               x10 : Bool;   // Direct output 1 via traversing block
               x11 : Bool;   // Direct output 2 via traversing block
               x12 : Bool;   // Fixed stop reached
               x13 : Bool;   // Fixed stop clamping torque reached
               x14 : Bool;   // Travel to fixed stop active
               x15 : Bool;   // Traversing command active
               x0 : Bool;   // Tracking mode active
               x1 : Bool;   // Velocity limit active
               x2 : Bool;   // Setpoint available
               x3 : Bool;   // Printing mark outside outer window
               x4 : Bool;   // Axis moves forwards
               x5 : Bool;   // Axis moves backwards
               x6 : Bool;   // Software limit switch minus reached
               x7 : Bool;   // Software limit switch plus reached
            END_STRUCT;
            dFDB_TARGET : DInt;   // R2060[5].Feedback target
            dXIST_A : DInt;   // R2521[0].Actual position value
            dNIST_B : DInt;   // R63.Actual speed value
            iFAULT_CODE : Int;   // R2131.Actual fault code
            iWARN_CODE : Int;   // R2132.Actual alarm code
            iUser : Int;
         END_STRUCT;
         tW : Struct   // WRITE
            tSTW1 : Struct   // CONTROL WORD 1
               x8 : Bool;   // P2589.EPOS jog 1 signal source
               x9 : Bool;   // P2590.EPOS jog 2 signal source
               x10 : Bool;   // P854[0].Control by PLC
               x11 : Bool;   // P2595.EPOS referencing start
               x12 : Bool;   // Reserved
               x13 : Bool;   // P2633.EPOS external block change
               x14 : Bool;   // Reserved
               x15 : Bool;   // P855[0] Brake release
               x0 : Bool;   // P840[0].ON/OFF
               x1 : Bool;   // P844[0].OFF2
               x2 : Bool;   // P848[0].OFF3
               x3 : Bool;   // P852[0].Enable operation
               x4 : Bool;   // P2641.EPOS abort traversing task
               x5 : Bool;   // P2640.EPOS intermediate STOP
               x6 : Bool;   // P2631.EPOS activate traversing task
               x7 : Bool;   // P2103.Acknowledge faults
            END_STRUCT;
            tPOS_STW1 : Struct   // POSITIONER CONTROL WORD 2
               x8 : Bool;   // P2648.EPOS direct setpoint input/MDI positioning type
               x9 : Bool;   // P2651.EPOS direct setpoint input/MDI direction selection positive
               x10 : Bool;   // P2652.EPOS direct setpoint input/MDI direction selection negative
               x11 : Bool;   // Reserved
               x12 : Bool;   // P2649.EPOS direct setpoint input/MDI transfer type selection
               x13 : Bool;   // Reserved
               x14 : Bool;   // P2653.EPOS direct setpoint input/MDI setting-up selection
               x15 : Bool;   // P2647.EPOS direct setpoint input/MDI selection
               x0 : Bool;   // P2525.EPOS traversing block selection, bit 0
               x1 : Bool;   // P2526.EPOS traversing block selection, bit 1
               x2 : Bool;   // P2527.EPOS traversing block selection, bit 2
               x3 : Bool;   // P2528.EPOS traversing block selection, bit 3
               x4 : Bool;   // P2529.EPOS traversing block selection, bit 4
               x5 : Bool;   // P2530.EPOS traversing block selection, bit 5
               x6 : Bool;   // Reserved
               x7 : Bool;   // Reserved
            END_STRUCT;
            tPOS_STW2 : Struct   // POSITIONER CONTROL WORD 3
               x8 : Bool;   // P2597.EPOS referencing type selection
               x9 : Bool;   // P2604.EPOS search for reference, start direction
               x10 : Bool;   // P2510.LR selecting measuring probe evaluation
               x11 : Bool;   // P2511.LR measuring probe evaluation edge
               x12 : Bool;   // Reserved
               x13 : Bool;   // Reserved
               x14 : Bool;   // P2582.EPOS software limit switch activation
               x15 : Bool;   // P2568.EPOS STOP cam activation
               x0 : Bool;   // P2655.EPOS select tracking mode
               x1 : Bool;   // P2596.EPOS set reference point
               x2 : Bool;   // P2612.EPOS search for reference cam
               x3 : Bool;   // Reserved
               x4 : Bool;   // Reserved
               x5 : Bool;   // P2591.EPOS jogging incremental
               x6 : Bool;   // Reserved
               x7 : Bool;   // Reserved
            END_STRUCT;
            iSTW2 : Int;   // P2045.CONTROL WORD 4
            iOVERRIDE : Int;   // P2646.Override % [0-16384]
            dMDI_TARPOS : DInt;   // P2642.Target position for MDI
            dMDI_VELOCITY : DInt;   // P2643.Speed reference for MDI
            iMDI_ACC : Int;   // P2644.Acceleration ramp % for MDI [0-16384]
            iMDI_DEC : Int;   // P2645.Deceleration ramp % for MDI [0-16384]
            iUser : Int;
         END_STRUCT;
      END_STRUCT;
   END_VAR
   VAR_TEMP
      TMP_dOldValue_AR1 : DInt;
      TMP_dOldValue_AR2 : DInt;
      TMP_x : Bool;
      TMP_i : Int;
      TMP_d : DInt;
      TMP_r : Real;
      TMP_a : ANY;
      TMP_dZero : DInt;
      TMP_xAlwaysON : Bool;
      TMP_rActualSpeed : Real;
      TMP_iAddressLength : Int;
      TMP_iRetVal : Int;
      TMP_dActualPosFiltered_cdeg : DInt;   // Actual position filtered [°/100]
      TMP_dActualPosMin_cdeg : DInt;   // Actual position minimum tollerance [°/100]
      TMP_dActualPosMax_cdeg : DInt;   // Actual position maximum tollerance [°/100]
   END_VAR
   VAR_TEMP   // added for the SCL form of the ladder/FBD networks
      _w1 : Bool;
      _w2 : Bool;
      _w3 : Bool;
      _w4 : Bool;
   END_VAR
BEGIN

REGION Network 1 (STL): Save AR1 & AR2 value
   //    TAR1
   //    T     #TMP_dOldValue_AR1
   //    TAR2
   //    T     #TMP_dOldValue_AR2
END_REGION

REGION Network 2: #####_COSTANTS_#####
END_REGION

REGION Network 3 (STL): Initializing
         SET;
         S     #TMP_xAlwaysON;

         L     DINT#0;
         T     #TMP_dZero;

         CALL  FILL
         ( BVAL    := #TMP_dZero,
           RET_VAL := #TMP_iRetVal,
           BLK     := #STC_tPZD_Pos.tR
         );

         CALL  FILL
         ( BVAL    := #TMP_dZero,
           RET_VAL := #TMP_iRetVal,
           BLK     := #STC_tMngSysReg
         );
END_REGION

REGION Network 4: #####_MOTOR_MODULE_#####
END_REGION

REGION Network 5 (STL): Check system data coerence
         L     #STC_tSYS_DATA.iIOAddress_MM;
         L     0;
         <I;
         L     10;
         JC    Err;

         L     #STC_tSYS_DATA.dMaxSpeed_rpm;
         L     DINT#0;
         <=D;
         L     11;
         JC    Err;

         L     #STC_tSYS_DATA.rK_rpm_grdMin;
         L     0.0;
         <=R;
         L     13;
         JC    Err;

         L     #STC_tSYS_DATA.rMaxAcc_deg_s2;
         L     0.0;
         <=R;
         L     14;
         JC    Err;

         L     #STC_tSYS_DATA.rMaxDec_deg_s2;
         L     0.0;
         <=R;
         L     15;
         JC    Err;
END_REGION

REGION Network 6: #####_MATCH_#####
END_REGION

REGION Network 7 (STL): Input copy
   // Compute destination position
         L;
         LAR1;
   //byte 1 = 10h (FIXED for S7)
         L     B#16#10;
         T     B[AR1, P#0.0];
   //byte 2 = data type
         L     B#16#4;  //4 = word
         T     B[AR1, P#1.0];
   //byte 3 & 4 = number of element
         L     12;  //Production data
         T     W[AR1, P#2.0];
   //byte 5 & 6 = number of DB
         L     0;  //DB production data
         T     W[AR1, P#4.0];
   //byte 7 = memory area
         L     B#16#81;  //81h = I (Input)
         T     B[AR1, P#6.0];
   //byte 8 & 9 = address. Bit 0,1,2 of tenth byte is bit offset
   //byte 7 = address (high). Valid value = 0-7. Bit 3,4,5,6,7 always 0
         L     #STC_tSYS_DATA.iIOAddress_MM;  //Item size
         SLW   3;
         T     W[AR1, P#8.0];
         SRD   16;
         AW    16#0007;
         T     B[AR1, P#7.0];
END_REGION

REGION Network 8: #########################_POSITIONER_###########################
END_REGION

REGION Network 9: #####_MATCH_#####
END_REGION

REGION Network 10 (STL): Input copy
         CALL  BLKMOV
         ( SRCBLK  := #TMP_a,
           RET_VAL := #TMP_iRetVal,
           DSTBLK  := #STC_tPZD_Pos.tR
         );
END_REGION

REGION Network 11: Status signals
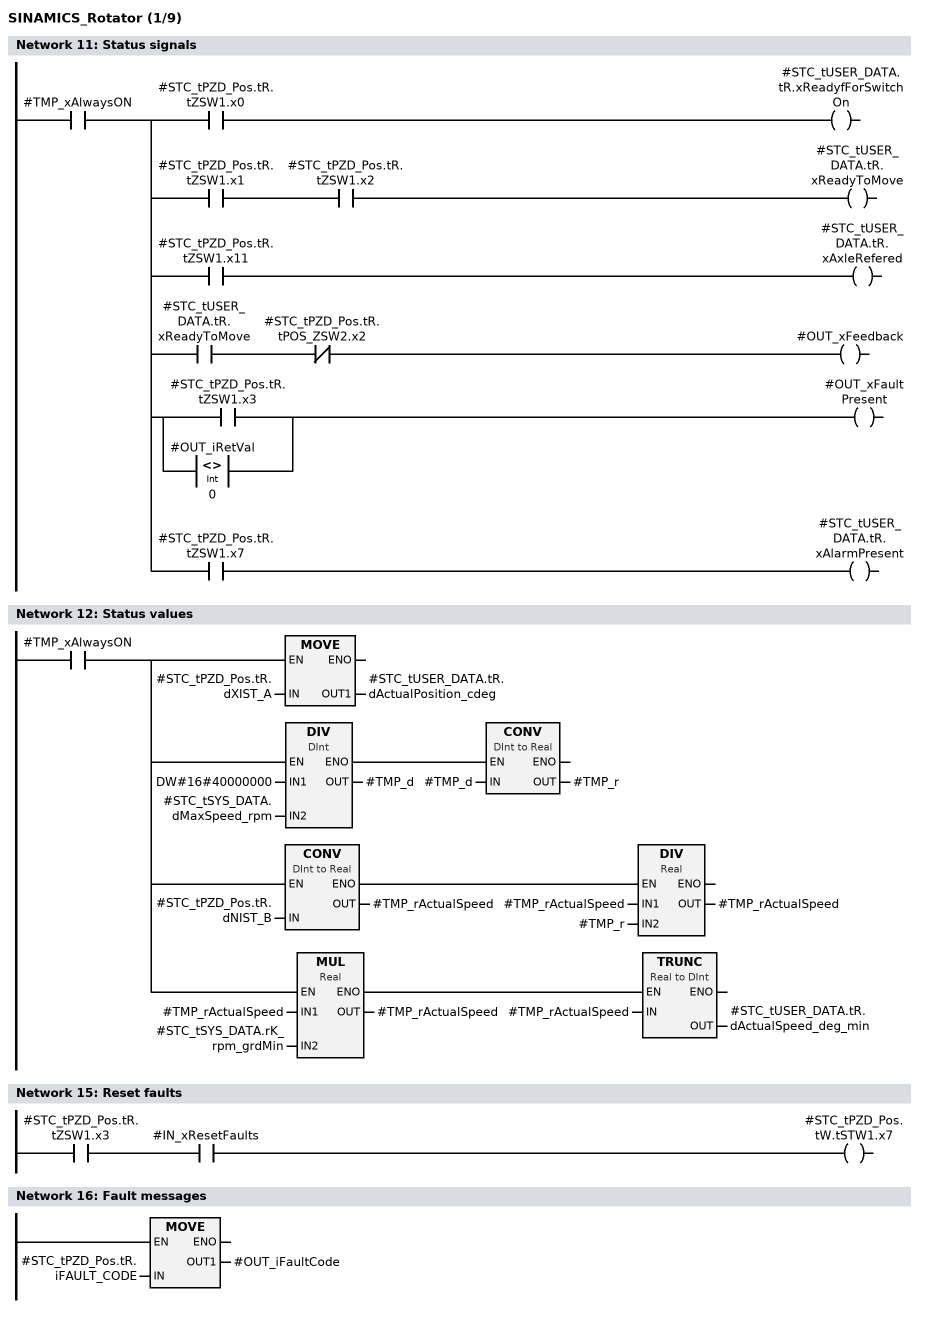
   RUNG wire#powerrail
      Contact( #TMP_xAlwaysON )
      wire#w1
      Contact( #STC_tPZD_Pos.tR.tZSW1.x0 )
      Coil( #STC_tUSER_DATA.tR.xReadyfForSwitchOn )
   END_RUNG
   RUNG wire#w1
      Contact( #STC_tPZD_Pos.tR.tZSW1.x1 )
      Contact( #STC_tPZD_Pos.tR.tZSW1.x2 )
      Coil( #STC_tUSER_DATA.tR.xReadyToMove )
   END_RUNG
   RUNG wire#w1
      Contact( #STC_tPZD_Pos.tR.tZSW1.x11 )
      Coil( #STC_tUSER_DATA.tR.xAxleRefered )
   END_RUNG
   RUNG wire#w1
      Contact( #STC_tUSER_DATA.tR.xReadyToMove )
      I_Contact( #STC_tPZD_Pos.tR.tPOS_ZSW2.x2 )
      Coil( #OUT_xFeedback )
   END_RUNG
   RUNG wire#w1
      Contact( #STC_tPZD_Pos.tR.tZSW1.x3 )
      wire#w2
      Coil( #OUT_xFaultPresent )
   END_RUNG
   RUNG wire#w1
      { S7_Templates := "SrcType := Int" } NE_Contact(in1 := #OUT_iRetVal, in2 := 0)
   END_RUNG wire#w2
   RUNG wire#w1
      Contact( #STC_tPZD_Pos.tR.tZSW1.x7 )
      Coil( #STC_tUSER_DATA.tR.xAlarmPresent )
   END_RUNG
   // the same network as SCL:
   #STC_tUSER_DATA.tR.xReadyfForSwitchOn := #TMP_xAlwaysON AND #STC_tPZD_Pos.tR.tZSW1.x0;
   #STC_tUSER_DATA.tR.xReadyToMove := #TMP_xAlwaysON AND #STC_tPZD_Pos.tR.tZSW1.x1 AND #STC_tPZD_Pos.tR.tZSW1.x2;
   #STC_tUSER_DATA.tR.xAxleRefered := #TMP_xAlwaysON AND #STC_tPZD_Pos.tR.tZSW1.x11;
   #OUT_xFeedback := #TMP_xAlwaysON AND #STC_tUSER_DATA.tR.xReadyToMove AND NOT #STC_tPZD_Pos.tR.tPOS_ZSW2.x2;
   #OUT_xFaultPresent := #TMP_xAlwaysON AND (#STC_tPZD_Pos.tR.tZSW1.x3 OR (#OUT_iRetVal <> 0));
   #STC_tUSER_DATA.tR.xAlarmPresent := #TMP_xAlwaysON AND #STC_tPZD_Pos.tR.tZSW1.x7;
END_REGION

REGION Network 12: Status values
   RUNG wire#powerrail
      Contact( #TMP_xAlwaysON )
      wire#w1
      { S7_GenerateENO := "TRUE" } Move(in := #STC_tPZD_Pos.tR.dXIST_A, out1 => #STC_tUSER_DATA.tR.dActualPosition_cdeg)
   END_RUNG
   RUNG wire#w1
      { S7_Templates := "SrcType := DInt"; S7_GenerateENO := "TRUE" } Div(in1 := DW#16#40000000, in2 := #STC_tSYS_DATA.dMaxSpeed_rpm, out => #TMP_d)
      { S7_Templates := "[SrcType := DInt, DestType := Real]"; S7_GenerateENO := "TRUE" } Convert(in := #TMP_d, out => #TMP_r)
   END_RUNG
   RUNG wire#w1
      { S7_Templates := "[SrcType := DInt, DestType := Real]"; S7_GenerateENO := "TRUE" } Convert(in := #STC_tPZD_Pos.tR.dNIST_B, out => #TMP_rActualSpeed)
      { S7_Templates := "SrcType := Real"; S7_GenerateENO := "TRUE" } Div(in1 := #TMP_rActualSpeed, in2 := #TMP_r, out => #TMP_rActualSpeed)
   END_RUNG
   RUNG wire#w1
      { S7_Templates := "SrcType := Real"; S7_GenerateENO := "TRUE" } Mul(in1 := #TMP_rActualSpeed, in2 := #STC_tSYS_DATA.rK_rpm_grdMin, out => #TMP_rActualSpeed)
      { S7_Templates := "[SrcType := Real, DestType := DInt]"; S7_GenerateENO := "TRUE" } Trunc(in := #TMP_rActualSpeed, out => #STC_tUSER_DATA.tR.dActualSpeed_deg_min)
   END_RUNG
   // the same network as SCL:
   // ENO of a box is taken as its EN; it also drops when the box reports an error
   IF #TMP_xAlwaysON THEN
       #STC_tUSER_DATA.tR.dActualPosition_cdeg := #STC_tPZD_Pos.tR.dXIST_A;
       #TMP_d := DW#16#40000000 / #STC_tSYS_DATA.dMaxSpeed_rpm;
       #TMP_r := DINT_TO_REAL(#TMP_d);
       #TMP_rActualSpeed := DINT_TO_REAL(#STC_tPZD_Pos.tR.dNIST_B);
       #TMP_rActualSpeed := #TMP_rActualSpeed / #TMP_r;
       #TMP_rActualSpeed := #TMP_rActualSpeed * #STC_tSYS_DATA.rK_rpm_grdMin;
       #STC_tUSER_DATA.tR.dActualSpeed_deg_min := TRUNC(#TMP_rActualSpeed);
   END_IF;
END_REGION

REGION Network 13: #####_STATUSES_#####
END_REGION

REGION Network 14: #####_ALARMS_#####
END_REGION

REGION Network 15: Reset faults
   RUNG wire#powerrail
      Contact( #STC_tPZD_Pos.tR.tZSW1.x3 )
      Contact( #IN_xResetFaults )
      Coil( #STC_tPZD_Pos.tW.tSTW1.x7 )
   END_RUNG
   // the same network as SCL:
   #STC_tPZD_Pos.tW.tSTW1.x7 := #STC_tPZD_Pos.tR.tZSW1.x3 AND #IN_xResetFaults;
END_REGION

REGION Network 16: Fault messages
   RUNG wire#powerrail
      { S7_GenerateENO := "TRUE" } Move(in := #STC_tPZD_Pos.tR.iFAULT_CODE, out1 => #OUT_iFaultCode)
   END_RUNG
   // the same network as SCL:
   #OUT_iFaultCode := #STC_tPZD_Pos.tR.iFAULT_CODE;
END_REGION

REGION Network 17: Alarm messages
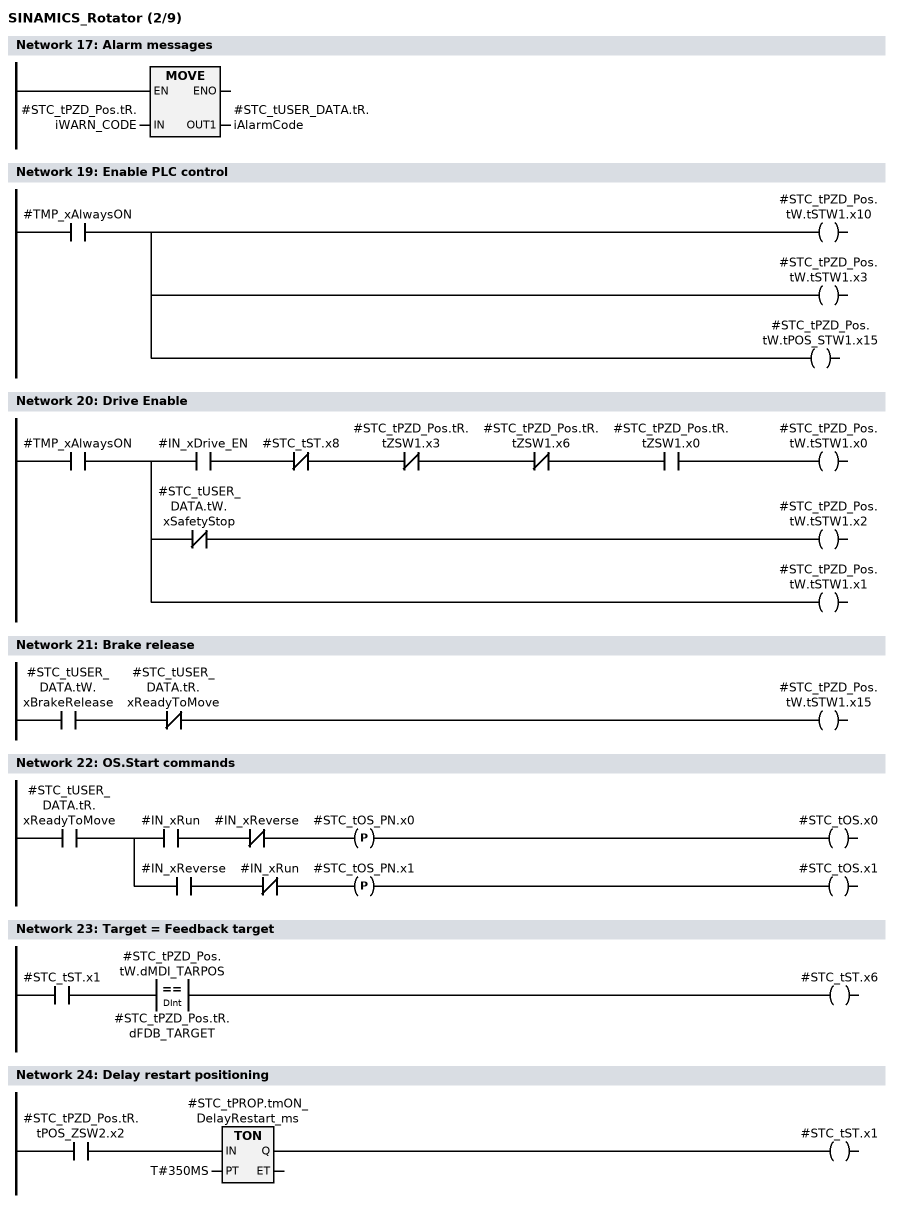
   RUNG wire#powerrail
      { S7_GenerateENO := "TRUE" } Move(in := #STC_tPZD_Pos.tR.iWARN_CODE, out1 => #STC_tUSER_DATA.tR.iAlarmCode)
   END_RUNG
   // the same network as SCL:
   #STC_tUSER_DATA.tR.iAlarmCode := #STC_tPZD_Pos.tR.iWARN_CODE;
END_REGION

REGION Network 18: #####_PHASES_&_LOGICS_#####
END_REGION

REGION Network 19: Enable PLC control
   RUNG wire#powerrail
      Contact( #TMP_xAlwaysON )
      wire#w1
      Coil( #STC_tPZD_Pos.tW.tSTW1.x10 )
   END_RUNG
   RUNG wire#w1
      Coil( #STC_tPZD_Pos.tW.tSTW1.x3 )
   END_RUNG
   RUNG wire#w1
      Coil( #STC_tPZD_Pos.tW.tPOS_STW1.x15 )
   END_RUNG
   // the same network as SCL:
   #STC_tPZD_Pos.tW.tSTW1.x10 := #TMP_xAlwaysON;
   #STC_tPZD_Pos.tW.tSTW1.x3 := #TMP_xAlwaysON;
   #STC_tPZD_Pos.tW.tPOS_STW1.x15 := #TMP_xAlwaysON;
END_REGION

REGION Network 20: Drive Enable
   RUNG wire#powerrail
      Contact( #TMP_xAlwaysON )
      wire#w1
      Contact( #IN_xDrive_EN )
      I_Contact( #STC_tST.x8 )
      I_Contact( #STC_tPZD_Pos.tR.tZSW1.x3 )
      I_Contact( #STC_tPZD_Pos.tR.tZSW1.x6 )
      Contact( #STC_tPZD_Pos.tR.tZSW1.x0 )
      Coil( #STC_tPZD_Pos.tW.tSTW1.x0 )
   END_RUNG
   RUNG wire#w1
      I_Contact( #STC_tUSER_DATA.tW.xSafetyStop )
      Coil( #STC_tPZD_Pos.tW.tSTW1.x2 )
   END_RUNG
   RUNG wire#w1
      Coil( #STC_tPZD_Pos.tW.tSTW1.x1 )
   END_RUNG
   // the same network as SCL:
   #STC_tPZD_Pos.tW.tSTW1.x0 := #TMP_xAlwaysON AND #IN_xDrive_EN AND NOT #STC_tST.x8 AND NOT #STC_tPZD_Pos.tR.tZSW1.x3 AND NOT #STC_tPZD_Pos.tR.tZSW1.x6 AND #STC_tPZD_Pos.tR.tZSW1.x0;
   #STC_tPZD_Pos.tW.tSTW1.x2 := #TMP_xAlwaysON AND NOT #STC_tUSER_DATA.tW.xSafetyStop;
   #STC_tPZD_Pos.tW.tSTW1.x1 := #TMP_xAlwaysON;
END_REGION

REGION Network 21: Brake release
   RUNG wire#powerrail
      Contact( #STC_tUSER_DATA.tW.xBrakeRelease )
      I_Contact( #STC_tUSER_DATA.tR.xReadyToMove )
      Coil( #STC_tPZD_Pos.tW.tSTW1.x15 )
   END_RUNG
   // the same network as SCL:
   #STC_tPZD_Pos.tW.tSTW1.x15 := #STC_tUSER_DATA.tW.xBrakeRelease AND NOT #STC_tUSER_DATA.tR.xReadyToMove;
END_REGION

REGION Network 22: OS.Start commands
   RUNG wire#powerrail
      Contact( #STC_tUSER_DATA.tR.xReadyToMove )
      wire#w1
      Contact( #IN_xRun )
      I_Contact( #IN_xReverse )
      P_Trig( #STC_tOS_PN.x0 )
      Coil( #STC_tOS.x0 )
   END_RUNG
   RUNG wire#w1
      Contact( #IN_xReverse )
      I_Contact( #IN_xRun )
      P_Trig( #STC_tOS_PN.x1 )
      Coil( #STC_tOS.x1 )
   END_RUNG
   // the same network as SCL:
   #_w1 := #STC_tUSER_DATA.tR.xReadyToMove AND #IN_xRun AND NOT #IN_xReverse;
   #_w2 := #_w1 AND NOT #STC_tOS_PN.x0;   // rising edge
   #STC_tOS_PN.x0 := #_w1;
   #STC_tOS.x0 := #_w2;
   #_w3 := #STC_tUSER_DATA.tR.xReadyToMove AND #IN_xReverse AND NOT #IN_xRun;
   #_w4 := #_w3 AND NOT #STC_tOS_PN.x1;   // rising edge
   #STC_tOS_PN.x1 := #_w3;
   #STC_tOS.x1 := #_w4;
END_REGION

REGION Network 23: Target = Feedback target
   RUNG wire#powerrail
      Contact( #STC_tST.x1 )
      { S7_Templates := "SrcType := DInt" } EQ_Contact(in1 := #STC_tPZD_Pos.tW.dMDI_TARPOS, in2 := #STC_tPZD_Pos.tR.dFDB_TARGET)
      Coil( #STC_tST.x6 )
   END_RUNG
   // the same network as SCL:
   #STC_tST.x6 := #STC_tST.x1 AND (#STC_tPZD_Pos.tW.dMDI_TARPOS = #STC_tPZD_Pos.tR.dFDB_TARGET);
END_REGION

REGION Network 24: Delay restart positioning
   #STC_tPROP.tmON_DelayRestart_ms.TON(IN := #STC_tPZD_Pos.tR.tPOS_ZSW2.x2, PT := T#350MS);
   #STC_tST.x1 := #STC_tPROP.tmON_DelayRestart_ms.Q;
END_REGION

REGION Network 25: Positioning request
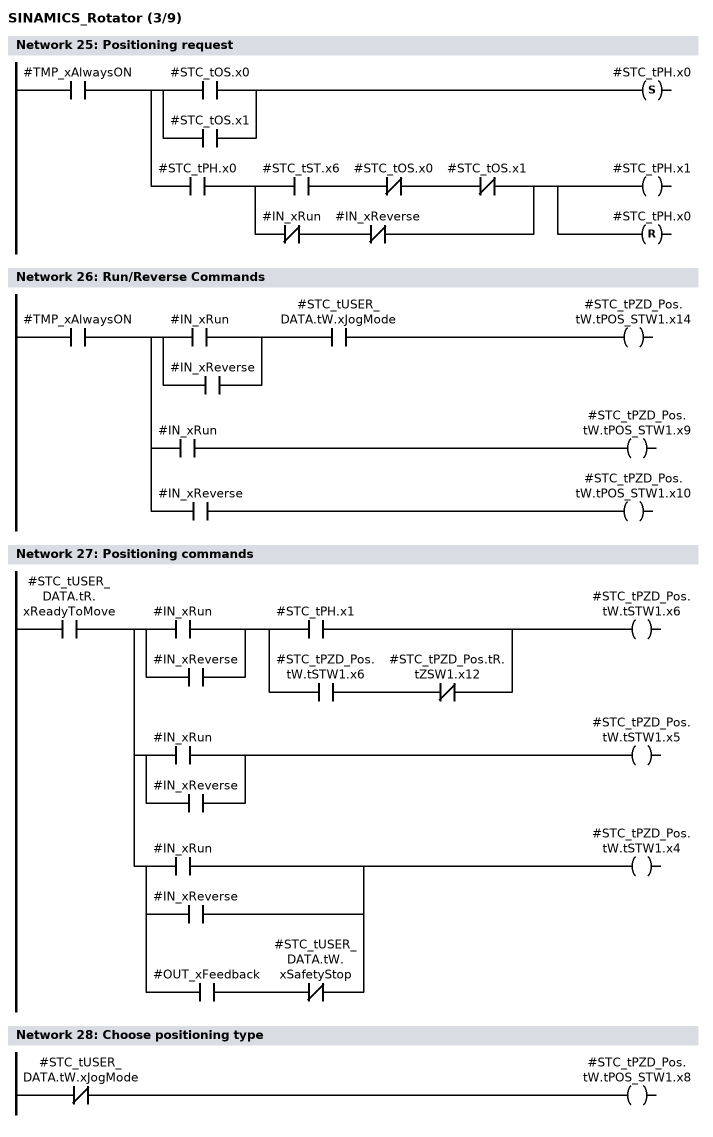
   RUNG wire#powerrail
      Contact( #TMP_xAlwaysON )
      wire#w1
      Contact( #STC_tOS.x0 )
      wire#w2
      S_Coil( #STC_tPH.x0 )
   END_RUNG
   RUNG wire#w1
      Contact( #STC_tOS.x1 )
   END_RUNG wire#w2
   RUNG wire#w1
      Contact( #STC_tPH.x0 )
      wire#w3
      Contact( #STC_tST.x6 )
      I_Contact( #STC_tOS.x0 )
      I_Contact( #STC_tOS.x1 )
      wire#w4
      Coil( #STC_tPH.x1 )
   END_RUNG
   RUNG wire#w3
      I_Contact( #IN_xRun )
      I_Contact( #IN_xReverse )
   END_RUNG wire#w4
   RUNG wire#w4
      R_Coil( #STC_tPH.x0 )
   END_RUNG
   // the same network as SCL:
   IF #TMP_xAlwaysON AND (#STC_tOS.x0 OR #STC_tOS.x1) THEN #STC_tPH.x0 := TRUE; END_IF;
   #STC_tPH.x1 := #TMP_xAlwaysON AND #STC_tPH.x0 AND ((#STC_tST.x6 AND NOT #STC_tOS.x0 AND NOT #STC_tOS.x1) OR (NOT #IN_xRun AND NOT #IN_xReverse));
   IF #STC_tPH.x1 THEN #STC_tPH.x0 := FALSE; END_IF;
END_REGION

REGION Network 26: Run/Reverse Commands
   RUNG wire#powerrail
      Contact( #TMP_xAlwaysON )
      wire#w1
      Contact( #IN_xRun )
      wire#w2
      Contact( #STC_tUSER_DATA.tW.xJogMode )
      Coil( #STC_tPZD_Pos.tW.tPOS_STW1.x14 )
   END_RUNG
   RUNG wire#w1
      Contact( #IN_xReverse )
   END_RUNG wire#w2
   RUNG wire#w1
      Contact( #IN_xRun )
      Coil( #STC_tPZD_Pos.tW.tPOS_STW1.x9 )
   END_RUNG
   RUNG wire#w1
      Contact( #IN_xReverse )
      Coil( #STC_tPZD_Pos.tW.tPOS_STW1.x10 )
   END_RUNG
   // the same network as SCL:
   #STC_tPZD_Pos.tW.tPOS_STW1.x14 := #TMP_xAlwaysON AND (#IN_xRun OR #IN_xReverse) AND #STC_tUSER_DATA.tW.xJogMode;
   #STC_tPZD_Pos.tW.tPOS_STW1.x9 := #TMP_xAlwaysON AND #IN_xRun;
   #STC_tPZD_Pos.tW.tPOS_STW1.x10 := #TMP_xAlwaysON AND #IN_xReverse;
END_REGION

REGION Network 27: Positioning commands
   RUNG wire#powerrail
      Contact( #STC_tUSER_DATA.tR.xReadyToMove )
      wire#w1
      Contact( #IN_xRun )
      wire#w2
      Contact( #STC_tPH.x1 )
      wire#w3
      Coil( #STC_tPZD_Pos.tW.tSTW1.x6 )
   END_RUNG
   RUNG wire#w1
      Contact( #IN_xReverse )
   END_RUNG wire#w2
   RUNG wire#w2
      Contact( #STC_tPZD_Pos.tW.tSTW1.x6 )
      I_Contact( #STC_tPZD_Pos.tR.tZSW1.x12 )
   END_RUNG wire#w3
   RUNG wire#w1
      Contact( #IN_xRun )
      wire#w4
      Coil( #STC_tPZD_Pos.tW.tSTW1.x5 )
   END_RUNG
   RUNG wire#w1
      Contact( #IN_xReverse )
   END_RUNG wire#w4
   RUNG wire#w1
      Contact( #IN_xRun )
      wire#w5
      Coil( #STC_tPZD_Pos.tW.tSTW1.x4 )
   END_RUNG
   RUNG wire#w1
      Contact( #IN_xReverse )
   END_RUNG wire#w5
   RUNG wire#w1
      Contact( #OUT_xFeedback )
      I_Contact( #STC_tUSER_DATA.tW.xSafetyStop )
   END_RUNG wire#w5
   // the same network as SCL:
   #STC_tPZD_Pos.tW.tSTW1.x6 := #STC_tUSER_DATA.tR.xReadyToMove AND (#IN_xRun OR #IN_xReverse) AND (#STC_tPH.x1 OR (#STC_tPZD_Pos.tW.tSTW1.x6 AND NOT #STC_tPZD_Pos.tR.tZSW1.x12));
   #STC_tPZD_Pos.tW.tSTW1.x5 := #STC_tUSER_DATA.tR.xReadyToMove AND (#IN_xRun OR #IN_xReverse);
   #STC_tPZD_Pos.tW.tSTW1.x4 := #STC_tUSER_DATA.tR.xReadyToMove AND (#IN_xRun OR #IN_xReverse OR (#OUT_xFeedback AND NOT #STC_tUSER_DATA.tW.xSafetyStop));
END_REGION

REGION Network 28: Choose positioning type
   RUNG wire#powerrail
      I_Contact( #STC_tUSER_DATA.tW.xJogMode )
      Coil( #STC_tPZD_Pos.tW.tPOS_STW1.x8 )
   END_RUNG
   // the same network as SCL:
   #STC_tPZD_Pos.tW.tPOS_STW1.x8 := NOT #STC_tUSER_DATA.tW.xJogMode;
END_REGION

REGION Network 29: Positioning reached
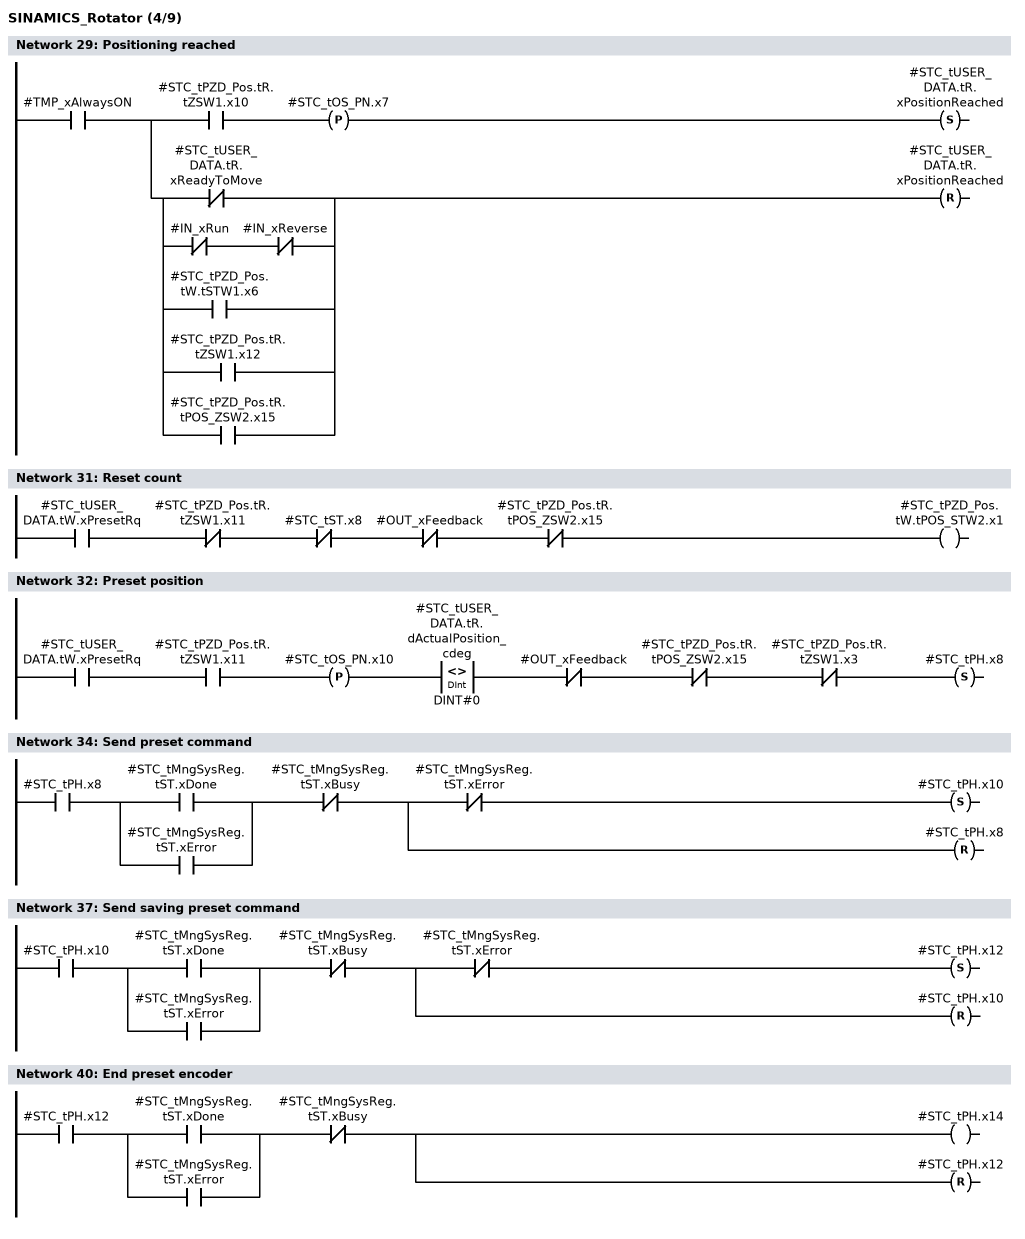
   RUNG wire#powerrail
      Contact( #TMP_xAlwaysON )
      wire#w1
      Contact( #STC_tPZD_Pos.tR.tZSW1.x10 )
      P_Trig( #STC_tOS_PN.x7 )
      S_Coil( #STC_tUSER_DATA.tR.xPositionReached )
   END_RUNG
   RUNG wire#w1
      I_Contact( #STC_tUSER_DATA.tR.xReadyToMove )
      wire#w2
      R_Coil( #STC_tUSER_DATA.tR.xPositionReached )
   END_RUNG
   RUNG wire#w1
      I_Contact( #IN_xRun )
      I_Contact( #IN_xReverse )
   END_RUNG wire#w2
   RUNG wire#w1
      Contact( #STC_tPZD_Pos.tW.tSTW1.x6 )
   END_RUNG wire#w2
   RUNG wire#w1
      Contact( #STC_tPZD_Pos.tR.tZSW1.x12 )
   END_RUNG wire#w2
   RUNG wire#w1
      Contact( #STC_tPZD_Pos.tR.tPOS_ZSW2.x15 )
   END_RUNG wire#w2
   // the same network as SCL:
   #_w1 := #TMP_xAlwaysON AND #STC_tPZD_Pos.tR.tZSW1.x10;
   #_w2 := #_w1 AND NOT #STC_tOS_PN.x7;   // rising edge
   #STC_tOS_PN.x7 := #_w1;
   IF #_w2 THEN #STC_tUSER_DATA.tR.xPositionReached := TRUE; END_IF;
   IF #TMP_xAlwaysON AND (NOT #STC_tUSER_DATA.tR.xReadyToMove OR (NOT #IN_xRun AND NOT #IN_xReverse) OR #STC_tPZD_Pos.tW.tSTW1.x6 OR #STC_tPZD_Pos.tR.tZSW1.x12 OR #STC_tPZD_Pos.tR.tPOS_ZSW2.x15) THEN
       #STC_tUSER_DATA.tR.xPositionReached := FALSE;
   END_IF;
END_REGION

REGION Network 30: #####_PRESET_ACTUAL_POSITION_#####
END_REGION

REGION Network 31: Reset count
   RUNG wire#powerrail
      Contact( #STC_tUSER_DATA.tW.xPresetRq )
      I_Contact( #STC_tPZD_Pos.tR.tZSW1.x11 )
      I_Contact( #STC_tST.x8 )
      I_Contact( #OUT_xFeedback )
      I_Contact( #STC_tPZD_Pos.tR.tPOS_ZSW2.x15 )
      Coil( #STC_tPZD_Pos.tW.tPOS_STW2.x1 )
   END_RUNG
   // the same network as SCL:
   #STC_tPZD_Pos.tW.tPOS_STW2.x1 := #STC_tUSER_DATA.tW.xPresetRq AND NOT #STC_tPZD_Pos.tR.tZSW1.x11 AND NOT #STC_tST.x8 AND NOT #OUT_xFeedback AND NOT #STC_tPZD_Pos.tR.tPOS_ZSW2.x15;
END_REGION

REGION Network 32: Preset position
   RUNG wire#powerrail
      Contact( #STC_tUSER_DATA.tW.xPresetRq )
      Contact( #STC_tPZD_Pos.tR.tZSW1.x11 )
      P_Trig( #STC_tOS_PN.x10 )
      { S7_Templates := "SrcType := DInt" } NE_Contact(in1 := #STC_tUSER_DATA.tR.dActualPosition_cdeg, in2 := DINT#0)
      I_Contact( #OUT_xFeedback )
      I_Contact( #STC_tPZD_Pos.tR.tPOS_ZSW2.x15 )
      I_Contact( #STC_tPZD_Pos.tR.tZSW1.x3 )
      S_Coil( #STC_tPH.x8 )
   END_RUNG
   // the same network as SCL:
   #_w1 := #STC_tUSER_DATA.tW.xPresetRq AND #STC_tPZD_Pos.tR.tZSW1.x11;
   #_w2 := #_w1 AND NOT #STC_tOS_PN.x10;   // rising edge
   #STC_tOS_PN.x10 := #_w1;
   IF #_w2 AND (#STC_tUSER_DATA.tR.dActualPosition_cdeg <> DINT#0) AND NOT #OUT_xFeedback AND NOT #STC_tPZD_Pos.tR.tPOS_ZSW2.x15 AND NOT #STC_tPZD_Pos.tR.tZSW1.x3 THEN
       #STC_tPH.x8 := TRUE;
   END_IF;
END_REGION

REGION Network 33 (STL): Send encoder value
         A     #STC_tPH.x8;
         JCN   PrE0;
         =     #STC_tMngSysReg.tST.xWrite_Request;

         L     #STC_tSYS_DATA.iPosPZD_MM;
         +     10;
         SLW   8;
         L     W#16#2;
         OW;
         T     #STC_tMngSysReg.tDATA.wRequest_refere_RequestID;
         L     #STC_tSYS_DATA.iPosPZD_MM;
         SLW   8;
         L     W#16#1;
         OW;
         T     #STC_tMngSysReg.tDATA.wAxis_NoOfParameters;
         L     W#16#1001;
         T     #STC_tMngSysReg.tDATA.wAttribute_NoOfElements;
         L     2599;
         T     #STC_tMngSysReg.tDATA.iParameter_number;
         L     W#16#0;
         T     #STC_tMngSysReg.tDATA.wSubindex;
         L     W#16#4301;
         T     #STC_tMngSysReg.tDATA.wFormat_NoOfValue;
         L     #STC_tSYS_DATA.iDiagAddress;
         T     #STC_tMngSysReg.tST.ID;
         L     47;
         T     #STC_tMngSysReg.tST.dINDEX;
         L     16;
         T     #STC_tMngSysReg.tST.uiLEN;

         L     DINT#0;
         T     #STC_tMngSysReg.tDATA.dwRegisterValue;

         CALL  #STC_tWriteRecord
         ( REQ    := #STC_tMngSysReg.tST.xWrite_Request,
           ID     := #STC_tMngSysReg.tST.ID,
           INDEX  := #STC_tMngSysReg.tST.dINDEX,
           LEN    := #STC_tMngSysReg.tST.uiLEN,
           DONE   := #STC_tMngSysReg.tST.xDone,
           BUSY   := #STC_tMngSysReg.tST.xBusy,
           ERROR  := #STC_tMngSysReg.tST.xError,
           STATUS := #STC_tMngSysReg.tST.dwSTATUS,
           RECORD := #STC_tMngSysReg.tDATA
         );
   PrE0: NOP   0;
END_REGION
